REGION Network 6
   RUNG wire#powerrail
      Contact( #iStop )
      Contact( #iRun )
      wire#w1
      R_Coil( #oON )
   END_RUNG
   RUNG wire#powerrail
      Contact( #oBlocked )
   END_RUNG wire#w1
   RUNG wire#w1
      R_Coil( #oBrake )
   END_RUNG
   RUNG wire#w1
      R_Coil( #oContactor )
   END_RUNG
   // the same network as SCL:
   IF (#iStop AND #iRun) OR #oBlocked THEN
       #oON := FALSE;
       #oBrake := FALSE;
       #oContactor := FALSE;
   END_IF;
END_REGION

REGION Network 7
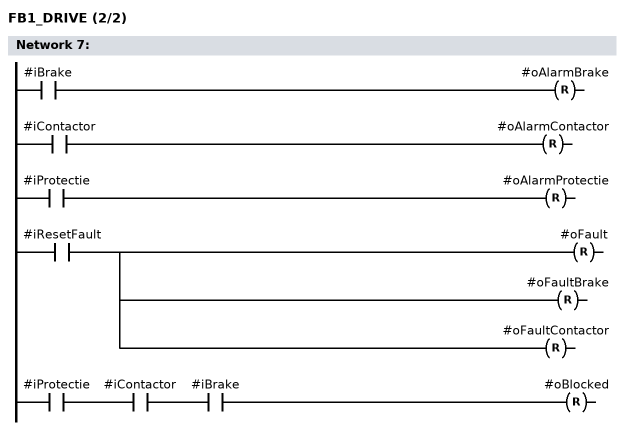
   RUNG wire#powerrail
      Contact( #iBrake )
      R_Coil( #oAlarmBrake )
   END_RUNG
   RUNG wire#powerrail
      Contact( #iContactor )
      R_Coil( #oAlarmContactor )
   END_RUNG
   RUNG wire#powerrail
      Contact( #iProtectie )
      R_Coil( #oAlarmProtectie )
   END_RUNG
   RUNG wire#powerrail
      Contact( #iResetFault )
      wire#w1
      R_Coil( #oFault )
   END_RUNG
   RUNG wire#w1
      R_Coil( #oFaultBrake )
   END_RUNG
   RUNG wire#w1
      R_Coil( #oFaultContactor )
   END_RUNG
   RUNG wire#powerrail
      Contact( #iProtectie )
      Contact( #iContactor )
      Contact( #iBrake )
      R_Coil( #oBlocked )
   END_RUNG
   // the same network as SCL:
   IF #iBrake THEN #oAlarmBrake := FALSE; END_IF;
   IF #iContactor THEN #oAlarmContactor := FALSE; END_IF;
   IF #iProtectie THEN #oAlarmProtectie := FALSE; END_IF;
   IF #iResetFault THEN
       #oFault := FALSE;
       #oFaultBrake := FALSE;
       #oFaultContactor := FALSE;
   END_IF;
   IF #iProtectie AND #iContactor AND #iBrake THEN #oBlocked := FALSE; END_IF;
END_REGION
END_FUNCTION_BLOCK

FUNCTION_BLOCK "FB_Pallet_Length"   // FB2, LAD
{ S7_Optimized_Access := 'TRUE' }
VERSION : 0.1
   VAR_INPUT
      iSQ_Pallet_Length : Bool;
      iConv_Speed : Int;
      Reset_Counter : Bool;
   END_VAR
   VAR_OUTPUT
      oPallet_Length : Int;
      oAlarm_Length : Bool;
   END_VAR
   VAR
      tSQ : Real;
      tMax : Time := T#20s;
      Pallet_count : Int;
      SQ_NOT : Bool;
      SQ_ON : Bool;
      Finished_counting : Bool;
   END_VAR
   VAR RETAIN
      Timer_ET : Time;
   END_VAR
   VAR
      Pallet_count_2 : Int;
      TON : TON_TIME;
   END_VAR
   VAR RETAIN
      CNT_PalletPass_2 : CTU_INT;
      CNT_PalletPass_1 : CTU_INT;
   END_VAR
   VAR_TEMP   // added for the SCL form of the ladder/FBD networks
      _w1 : Bool;
      _w2 : Bool;
   END_VAR
BEGIN

REGION Network 1
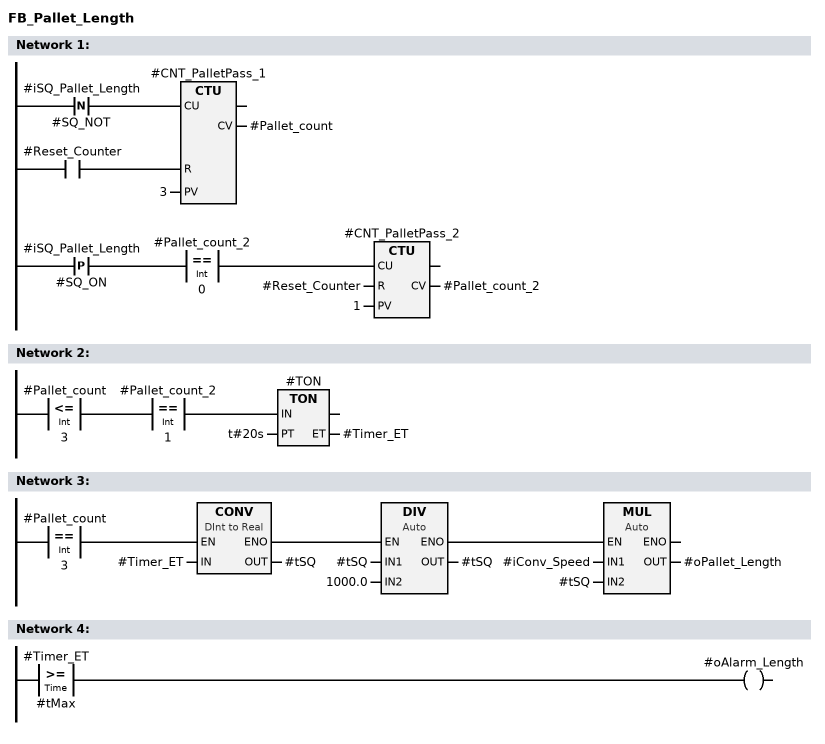
   #_w1 := NOT #iSQ_Pallet_Length AND #SQ_NOT;   // falling edge of #iSQ_Pallet_Length
   #SQ_NOT := #iSQ_Pallet_Length;
   #CNT_PalletPass_1(CU := #_w1, R := #Reset_Counter, PV := 3, CV => #Pallet_count);   // CTU
   #_w2 := #iSQ_Pallet_Length AND NOT #SQ_ON;   // rising edge of #iSQ_Pallet_Length
   #SQ_ON := #iSQ_Pallet_Length;
   #CNT_PalletPass_2(CU := #_w2 AND (#Pallet_count_2 = 0), R := #Reset_Counter, PV := 1, CV => #Pallet_count_2);   // CTU
END_REGION

REGION Network 2
   #TON(IN := (#Pallet_count <= 3) AND (#Pallet_count_2 = 1), PT := t#20s, ET => #Timer_ET);   // TON
END_REGION

REGION Network 3
   RUNG wire#powerrail
      { S7_Templates := "SrcType := Int" } EQ_Contact(in1 := #Pallet_count, in2 := 3)
      { S7_Templates := "[SrcType := DInt, DestType := Real]" } Convert(in := #Timer_ET, out => #tSQ)
      Div(in1 := #tSQ, in2 := 1000.0, out => #tSQ)
      Mul(in1 := #iConv_Speed, in2 := #tSQ, out => #oPallet_Length)
   END_RUNG
   // the same network as SCL:
   IF #Pallet_count = 3 THEN
       #tSQ := DINT_TO_REAL(#Timer_ET);
       #tSQ := #tSQ / 1000.0;
       #oPallet_Length := #iConv_Speed * #tSQ;
   END_IF;
END_REGION

REGION Network 4
   RUNG wire#powerrail
      { S7_Templates := "SrcType := Time" } GE_Contact(in1 := #Timer_ET, in2 := #tMax)
      Coil( #oAlarm_Length )
   END_RUNG
   // the same network as SCL:
   #oAlarm_Length := #Timer_ET >= #tMax;
END_REGION
END_FUNCTION_BLOCK

FUNCTION_BLOCK "FB_DS_Check_Machine"   // FB3, LAD
{ S7_Optimized_Access := 'TRUE' }
VERSION : 0.1
   VAR_INPUT
      iAir : Bool;
      iProtectie_CD_Drive : Bool;
      iProtectie_DS_Drive : Bool;
      iCD_Drive_Fault : Bool;
      iDS_Drive_Fault : Bool;
      iDestacker_Wait_Position : Bool;
      iSoftStarter_S1 : Bool;
      iSoftStarter_S2 : Bool;
   END_VAR
   VAR_OUTPUT
      oDS_Checked : Bool;
      oCD_Drive_NOK : Bool;
      oDS_Drive_NOK : Bool;
      oAir_NOK : Bool;
      oPower_NOK : Bool;
      oDestacker_NOK : Bool;
   END_VAR
   VAR
      AIR_OK : Bool;
      POWER_OK : Bool;
      Destacker_Wait_Position : Bool;
      CD_DRIVE_OK : Bool;
      DS_DRIVE_OK : Bool;
   END_VAR
BEGIN

REGION Network 1
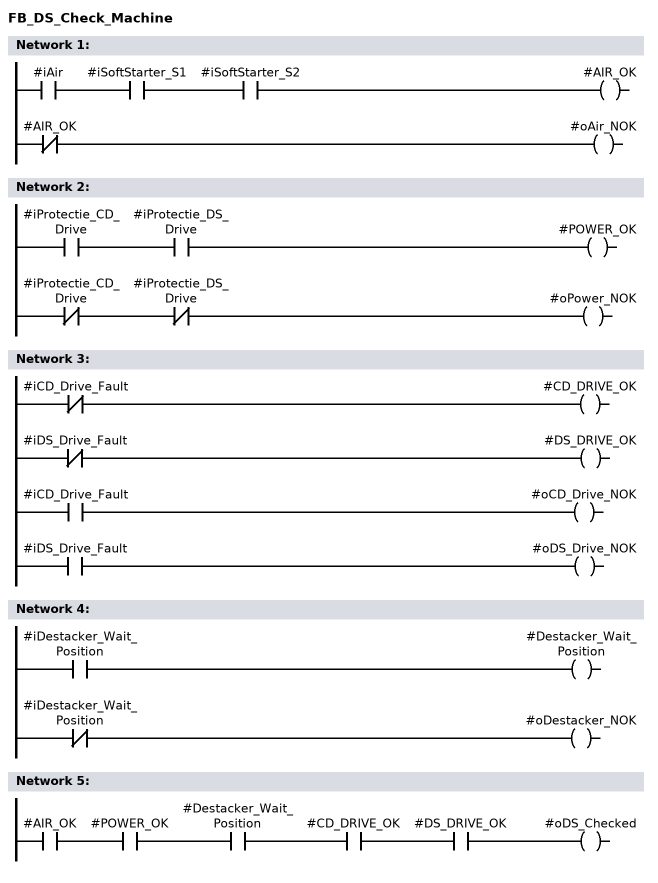
   RUNG wire#powerrail
      Contact( #iAir )
      Contact( #iSoftStarter_S1 )
      Contact( #iSoftStarter_S2 )
      Coil( #AIR_OK )
   END_RUNG
   RUNG wire#powerrail
      I_Contact( #AIR_OK )
      Coil( #oAir_NOK )
   END_RUNG
   // the same network as SCL:
   #AIR_OK := #iAir AND #iSoftStarter_S1 AND #iSoftStarter_S2;
   #oAir_NOK := NOT #AIR_OK;
END_REGION

REGION Network 2
   RUNG wire#powerrail
      Contact( #iProtectie_CD_Drive )
      Contact( #iProtectie_DS_Drive )
      Coil( #POWER_OK )
   END_RUNG
   RUNG wire#powerrail
      I_Contact( #iProtectie_CD_Drive )
      I_Contact( #iProtectie_DS_Drive )
      Coil( #oPower_NOK )
   END_RUNG
   // the same network as SCL:
   #POWER_OK := #iProtectie_CD_Drive AND #iProtectie_DS_Drive;
   #oPower_NOK := NOT #iProtectie_CD_Drive AND NOT #iProtectie_DS_Drive;
END_REGION

REGION Network 3
   RUNG wire#powerrail
      I_Contact( #iCD_Drive_Fault )
      Coil( #CD_DRIVE_OK )
   END_RUNG
   RUNG wire#powerrail
      I_Contact( #iDS_Drive_Fault )
      Coil( #DS_DRIVE_OK )
   END_RUNG
   RUNG wire#powerrail
      Contact( #iCD_Drive_Fault )
      Coil( #oCD_Drive_NOK )
   END_RUNG
   RUNG wire#powerrail
      Contact( #iDS_Drive_Fault )
      Coil( #oDS_Drive_NOK )
   END_RUNG
   // the same network as SCL:
   #CD_DRIVE_OK := NOT #iCD_Drive_Fault;
   #DS_DRIVE_OK := NOT #iDS_Drive_Fault;
   #oCD_Drive_NOK := #iCD_Drive_Fault;
   #oDS_Drive_NOK := #iDS_Drive_Fault;
END_REGION

REGION Network 4
   RUNG wire#powerrail
      Contact( #iDestacker_Wait_Position )
      Coil( #Destacker_Wait_Position )
   END_RUNG
   RUNG wire#powerrail
      I_Contact( #iDestacker_Wait_Position )
      Coil( #oDestacker_NOK )
   END_RUNG
   // the same network as SCL:
   #Destacker_Wait_Position := #iDestacker_Wait_Position;
   #oDestacker_NOK := NOT #iDestacker_Wait_Position;
END_REGION

REGION Network 5
   RUNG wire#powerrail
      Contact( #AIR_OK )
      Contact( #POWER_OK )
      Contact( #Destacker_Wait_Position )
      Contact( #CD_DRIVE_OK )
      Contact( #DS_DRIVE_OK )
      Coil( #oDS_Checked )
   END_RUNG
   // the same network as SCL:
   #oDS_Checked := #AIR_OK AND #POWER_OK AND #Destacker_Wait_Position AND #CD_DRIVE_OK AND #DS_DRIVE_OK;
END_REGION
END_FUNCTION_BLOCK

FUNCTION_BLOCK "FB_Init_S"   // FB4, LAD
TITLE = td -bitii de comenzi locali (ex: #Comanda_Furca) trebuie pusi in OUT
{ S7_Optimized_Access := 'TRUE' }
VERSION : 0.1
   VAR_INPUT
      DRV : "Bits_Stacker";
   END_VAR
   VAR
      Vertical : Bool;
      Furca : Bool;
      Comanda_Furca : Bool;
      Comanda_Vertical : Bool;
      InitReq : Bool;
      Init_OK : Bool;
      Alarm_Timeout_Vertical : Bool;
      Alarm_Timeout_Furca : Bool;
      "step" : USInt;
      Init_NotPossible : Bool;
      RstStack : Bool;
      Timer_Alarms : Array[0..1] of IEC_TIMER;
   END_VAR
   VAR_TEMP   // added for the SCL form of the ladder/FBD networks
      _w1 : Bool;
      _w2 : Bool;
   END_VAR
BEGIN

REGION Network 1: ini req
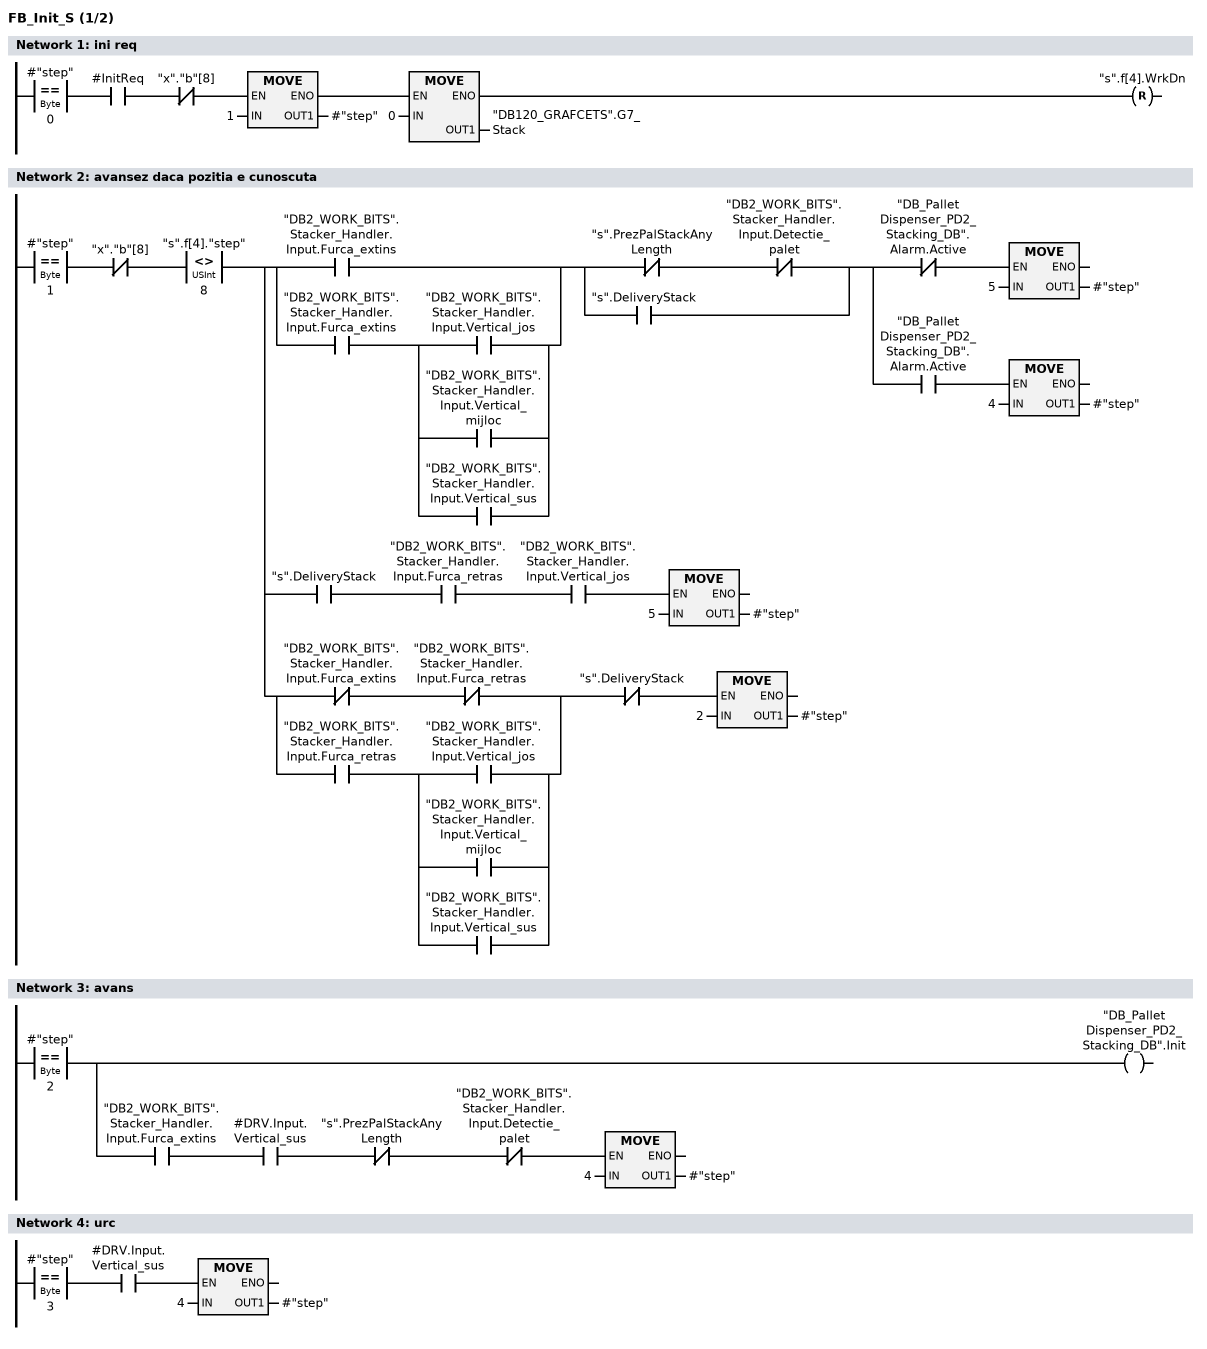
   RUNG wire#powerrail
      { S7_Templates := "SrcType := Byte" } EQ_Contact(in1 := #"step", in2 := 0)
      Contact( #InitReq )
      I_Contact( "x"."b"[8] )
      Move(in := 1, out1 => #"step")
      Move(in := 0, out1 => "DB120_GRAFCETS".G7_Stack)
      R_Coil( "s".f[4].WrkDn )
   END_RUNG
   // the same network as SCL:
   #_w1 := (#"step" = 0) AND #InitReq AND NOT "x"."b"[8];
   IF #_w1 THEN
       #"step" := 1;
       "DB120_GRAFCETS".G7_Stack := 0;
       "s".f[4].WrkDn := FALSE;
   END_IF;
END_REGION

REGION Network 2: avansez daca pozitia e cunoscuta
   RUNG wire#powerrail
      { S7_Templates := "SrcType := Byte" } EQ_Contact(in1 := #"step", in2 := 1)
      I_Contact( "x"."b"[8] )
      { S7_Templates := "SrcType := USInt" } NE_Contact(in1 := "s".f[4]."step", in2 := 8)
      wire#w1
      Contact( "DB2_WORK_BITS".Stacker_Handler.Input.Furca_extins )
      wire#w2
      I_Contact( "s".PrezPalStackAnyLength )
      I_Contact( "DB2_WORK_BITS".Stacker_Handler.Input.Detectie_palet )
      wire#w4
      I_Contact( "DB_PalletDispenser_PD2_Stacking_DB".Alarm.Active )
      Move(in := 5, out1 => #"step")
   END_RUNG
   RUNG wire#w1
      Contact( "DB2_WORK_BITS".Stacker_Handler.Input.Furca_extins )
      wire#w3
      Contact( "DB2_WORK_BITS".Stacker_Handler.Input.Vertical_jos )
   END_RUNG wire#w2
   RUNG wire#w3
      Contact( "DB2_WORK_BITS".Stacker_Handler.Input.Vertical_mijloc )
   END_RUNG wire#w2
   RUNG wire#w3
      Contact( "DB2_WORK_BITS".Stacker_Handler.Input.Vertical_sus )
   END_RUNG wire#w2
   RUNG wire#w2
      Contact( "s".DeliveryStack )
   END_RUNG wire#w4
   RUNG wire#w4
      Contact( "DB_PalletDispenser_PD2_Stacking_DB".Alarm.Active )
      Move(in := 4, out1 => #"step")
   END_RUNG
   RUNG wire#w1
      Contact( "s".DeliveryStack )
      Contact( "DB2_WORK_BITS".Stacker_Handler.Input.Furca_retras )
      Contact( "DB2_WORK_BITS".Stacker_Handler.Input.Vertical_jos )
      Move(in := 5, out1 => #"step")
   END_RUNG
   RUNG wire#w1
      I_Contact( "DB2_WORK_BITS".Stacker_Handler.Input.Furca_extins )
      I_Contact( "DB2_WORK_BITS".Stacker_Handler.Input.Furca_retras )
      wire#w5
      I_Contact( "s".DeliveryStack )
      Move(in := 2, out1 => #"step")
   END_RUNG
   RUNG wire#w1
      Contact( "DB2_WORK_BITS".Stacker_Handler.Input.Furca_retras )
      wire#w6
      Contact( "DB2_WORK_BITS".Stacker_Handler.Input.Vertical_jos )
   END_RUNG wire#w5
   RUNG wire#w6
      Contact( "DB2_WORK_BITS".Stacker_Handler.Input.Vertical_mijloc )
   END_RUNG wire#w5
   RUNG wire#w6
      Contact( "DB2_WORK_BITS".Stacker_Handler.Input.Vertical_sus )
   END_RUNG wire#w5
   // the same network as SCL:
   #_w1 := (#"step" = 1) AND NOT "x"."b"[8] AND ("s".f[4]."step" <> 8);
   #_w2 := #_w1 AND ("DB2_WORK_BITS".Stacker_Handler.Input.Furca_extins OR ("DB2_WORK_BITS".Stacker_Handler.Input.Furca_extins AND ("DB2_WORK_BITS".Stacker_Handler.Input.Vertical_jos OR "DB2_WORK_BITS".Stacker_Handler.Input.Vertical_mijloc OR "DB2_WORK_BITS".Stacker_Handler.Input.Vertical_sus))) AND ((NOT "s".PrezPalStackAnyLength AND NOT "DB2_WORK_BITS".Stacker_Handler.Input.Detectie_palet) OR "s".DeliveryStack);
   IF #_w2 AND NOT "DB_PalletDispenser_PD2_Stacking_DB".Alarm.Active THEN #"step" := 5; END_IF;
   IF #_w2 AND "DB_PalletDispenser_PD2_Stacking_DB".Alarm.Active THEN #"step" := 4; END_IF;
   IF #_w1 AND "s".DeliveryStack AND "DB2_WORK_BITS".Stacker_Handler.Input.Furca_retras AND "DB2_WORK_BITS".Stacker_Handler.Input.Vertical_jos THEN
       #"step" := 5;
   END_IF;
   IF #_w1 AND ((NOT "DB2_WORK_BITS".Stacker_Handler.Input.Furca_extins AND NOT "DB2_WORK_BITS".Stacker_Handler.Input.Furca_retras) OR ("DB2_WORK_BITS".Stacker_Handler.Input.Furca_retras AND ("DB2_WORK_BITS".Stacker_Handler.Input.Vertical_jos OR "DB2_WORK_BITS".Stacker_Handler.Input.Vertical_mijloc OR "DB2_WORK_BITS".Stacker_Handler.Input.Vertical_sus))) AND NOT "s".DeliveryStack THEN
       #"step" := 2;
   END_IF;
END_REGION

REGION Network 3: avans
   RUNG wire#powerrail
      { S7_Templates := "SrcType := Byte" } EQ_Contact(in1 := #"step", in2 := 2)
      wire#w1
      Coil( "DB_PalletDispenser_PD2_Stacking_DB".Init )
   END_RUNG
   RUNG wire#w1
      Contact( "DB2_WORK_BITS".Stacker_Handler.Input.Furca_extins )
      Contact( #DRV.Input.Vertical_sus )
      I_Contact( "s".PrezPalStackAnyLength )
      I_Contact( "DB2_WORK_BITS".Stacker_Handler.Input.Detectie_palet )
      Move(in := 4, out1 => #"step")
   END_RUNG
   // the same network as SCL:
   "DB_PalletDispenser_PD2_Stacking_DB".Init := #"step" = 2;
   IF "DB_PalletDispenser_PD2_Stacking_DB".Init AND "DB2_WORK_BITS".Stacker_Handler.Input.Furca_extins AND #DRV.Input.Vertical_sus AND NOT "s".PrezPalStackAnyLength AND NOT "DB2_WORK_BITS".Stacker_Handler.Input.Detectie_palet THEN
       #"step" := 4;
   END_IF;
END_REGION

REGION Network 4: urc
   RUNG wire#powerrail
      { S7_Templates := "SrcType := Byte" } EQ_Contact(in1 := #"step", in2 := 3)
      Contact( #DRV.Input.Vertical_sus )
      Move(in := 4, out1 => #"step")
   END_RUNG
   // the same network as SCL:
   IF (#"step" = 3) AND #DRV.Input.Vertical_sus THEN #"step" := 4; END_IF;
END_REGION

REGION Network 5: Reset FB stacker errors
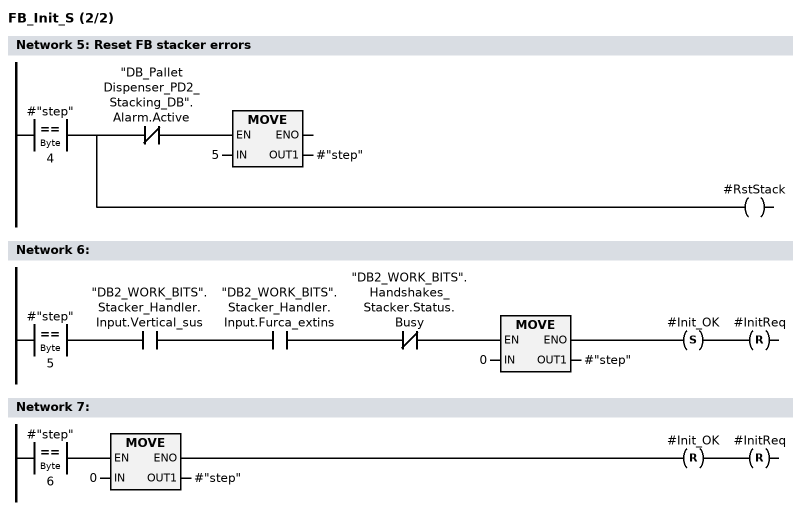
   RUNG wire#powerrail
      { S7_Templates := "SrcType := Byte" } EQ_Contact(in1 := #"step", in2 := 4)
      wire#w1
      I_Contact( "DB_PalletDispenser_PD2_Stacking_DB".Alarm.Active )
      Move(in := 5, out1 => #"step")
   END_RUNG
   RUNG wire#w1
      Coil( #RstStack )
   END_RUNG
   // the same network as SCL:
   #_w1 := #"step" = 4;
   IF #_w1 AND NOT "DB_PalletDispenser_PD2_Stacking_DB".Alarm.Active THEN #"step" := 5; END_IF;
   #RstStack := #_w1;
END_REGION

REGION Network 6
   RUNG wire#powerrail
      { S7_Templates := "SrcType := Byte" } EQ_Contact(in1 := #"step", in2 := 5)
      Contact( "DB2_WORK_BITS".Stacker_Handler.Input.Vertical_sus )
      Contact( "DB2_WORK_BITS".Stacker_Handler.Input.Furca_extins )
      I_Contact( "DB2_WORK_BITS".Handshakes_Stacker.Status.Busy )
      Move(in := 0, out1 => #"step")
      S_Coil( #Init_OK )
      R_Coil( #InitReq )
   END_RUNG
   // the same network as SCL:
   #_w1 := (#"step" = 5) AND "DB2_WORK_BITS".Stacker_Handler.Input.Vertical_sus AND "DB2_WORK_BITS".Stacker_Handler.Input.Furca_extins AND NOT "DB2_WORK_BITS".Handshakes_Stacker.Status.Busy;
   IF #_w1 THEN
       #"step" := 0;
       #Init_OK := TRUE;
       #InitReq := FALSE;
   END_IF;
END_REGION

REGION Network 7
   RUNG wire#powerrail
      { S7_Templates := "SrcType := Byte" } EQ_Contact(in1 := #"step", in2 := 6)
      Move(in := 0, out1 => #"step")
      R_Coil( #Init_OK )
      R_Coil( #InitReq )
   END_RUNG
   // the same network as SCL:
   #_w1 := #"step" = 6;
   IF #_w1 THEN
       #"step" := 0;
       #Init_OK := FALSE;
       #InitReq := FALSE;
   END_IF;
END_REGION
END_FUNCTION_BLOCK

FUNCTION_BLOCK "FB_Centrare"   // FB5, LAD
{ S7_Optimized_Access := 'TRUE' }
VERSION : 0.1
   VAR_INPUT
      Senzor_eliber : Bool;
      senzor_centr : Bool;
      step_st : USInt;
   END_VAR
   VAR_OUTPUT
      Comanda_centr : Bool;
      Comanda_eliber : Bool;
      stpo : USInt;
   END_VAR
   VAR_IN_OUT
      work : Bool;
   END_VAR
   VAR
      "step" : USInt;
      cmdav : Bool;
      cmdret : Bool;
      tmr : Array[1..3] of IEC_TIMER;
   END_VAR
   VAR_TEMP   // added for the SCL form of the ladder/FBD networks
      _w1 : Bool;
      _w2 : Bool;
   END_VAR
BEGIN

REGION Network 1
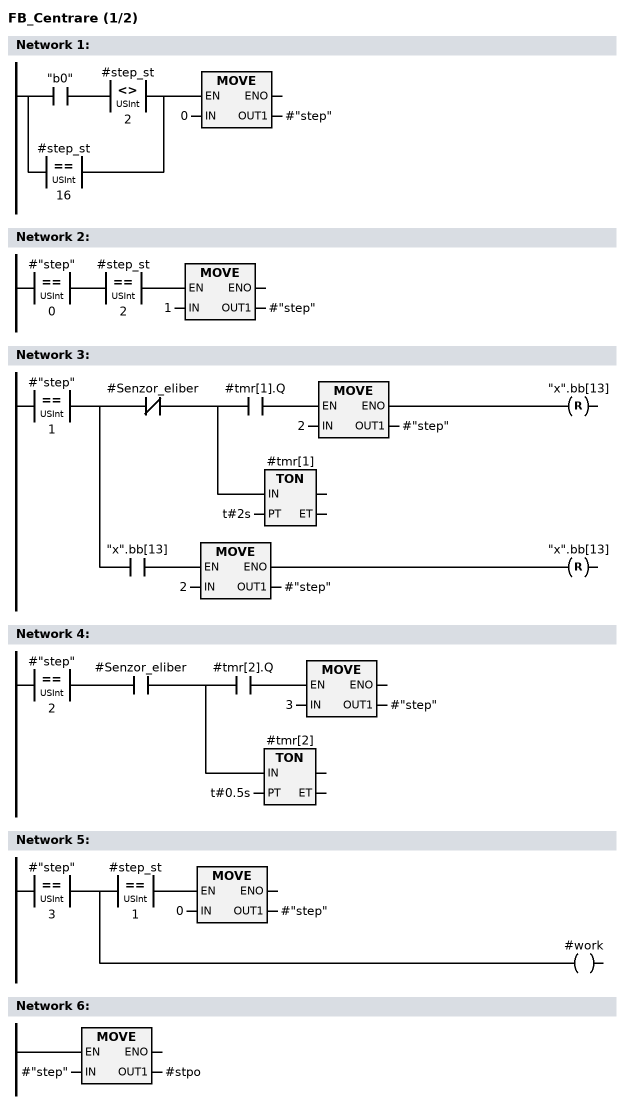
   RUNG wire#powerrail
      Contact( "b0" )
      { S7_Templates := "SrcType := USInt" } NE_Contact(in1 := #step_st, in2 := 2)
      wire#w1
      Move(in := 0, out1 => #"step")
   END_RUNG
   RUNG wire#powerrail
      { S7_Templates := "SrcType := USInt" } EQ_Contact(in1 := #step_st, in2 := 16)
   END_RUNG wire#w1
   // the same network as SCL:
   IF ("b0" AND (#step_st <> 2)) OR (#step_st = 16) THEN #"step" := 0; END_IF;
END_REGION

REGION Network 2
   RUNG wire#powerrail
      { S7_Templates := "SrcType := USInt" } EQ_Contact(in1 := #"step", in2 := 0)
      { S7_Templates := "SrcType := USInt" } EQ_Contact(in1 := #step_st, in2 := 2)
      Move(in := 1, out1 => #"step")
   END_RUNG
   // the same network as SCL:
   IF (#"step" = 0) AND (#step_st = 2) THEN #"step" := 1; END_IF;
END_REGION

REGION Network 3
   #_w1 := #"step" = 1;
   #_w2 := #_w1 AND NOT #Senzor_eliber;
   IF #_w2 AND #tmr[1].Q THEN
       #"step" := 2;
       "x".bb[13] := FALSE;
   END_IF;
   #tmr[1].TON(IN := #_w2, PT := t#2s);
   IF #_w1 AND "x".bb[13] THEN
       #"step" := 2;
       "x".bb[13] := FALSE;
   END_IF;
END_REGION

REGION Network 4
   #_w1 := (#"step" = 2) AND #Senzor_eliber;
   IF #_w1 AND #tmr[2].Q THEN #"step" := 3; END_IF;
   #tmr[2].TON(IN := #_w1, PT := t#0.5s);
END_REGION

REGION Network 5
   RUNG wire#powerrail
      { S7_Templates := "SrcType := USInt" } EQ_Contact(in1 := #"step", in2 := 3)
      wire#w1
      { S7_Templates := "SrcType := USInt" } EQ_Contact(in1 := #step_st, in2 := 1)
      Move(in := 0, out1 => #"step")
   END_RUNG
   RUNG wire#w1
      Coil( #work )
   END_RUNG
   // the same network as SCL:
   #_w1 := #"step" = 3;
   IF #_w1 AND (#step_st = 1) THEN #"step" := 0; END_IF;
   #work := #_w1;
END_REGION

REGION Network 6
   RUNG wire#powerrail
      Move(in := #"step", out1 => #stpo)
   END_RUNG
   // the same network as SCL:
   #stpo := #"step";
END_REGION

REGION Network 7: Apelare centror
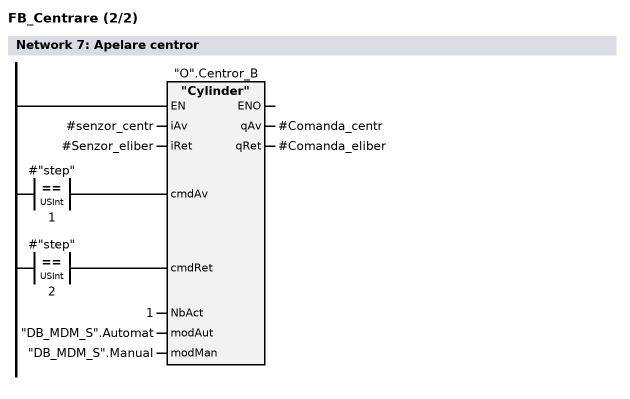
   RUNG wire#powerrail
      "O".Centror_B(cmdAv := wire#w1, cmdRet := wire#w2, iAv := #senzor_centr, iRet := #Senzor_eliber, NbAct := 1, modAut := "DB_MDM_S".Automat, modMan := "DB_MDM_S".Manual, qAv => #Comanda_centr, qRet => #Comanda_eliber)
   END_RUNG
   RUNG wire#powerrail
      { S7_Templates := "SrcType := USInt" } EQ_Contact(in1 := #"step", in2 := 1)
   END_RUNG wire#w1
   RUNG wire#powerrail
      { S7_Templates := "SrcType := USInt" } EQ_Contact(in1 := #"step", in2 := 2)
   END_RUNG wire#w2
   // the same network as SCL:
   "O".Centror_B(iAv := #senzor_centr,   // "Cylinder"
                 iRet := #Senzor_eliber,
                 cmdAv := #"step" = 1,
                 cmdRet := #"step" = 2,
                 NbAct := 1,
                 modAut := "DB_MDM_S".Automat,
                 modMan := "DB_MDM_S".Manual,
                 qAv => #Comanda_centr,
                 qRet => #Comanda_eliber);
END_REGION
END_FUNCTION_BLOCK

FUNCTION_BLOCK "sim"   // FB6, LAD
{ S7_Optimized_Access := 'TRUE' }
VERSION : 0.1
   VAR
      cen : "simCylinder";
      stH : "simCylinder";
      tct : IEC_TIMER;
      tct2 : Bool;
      tct1 : Bool;
      tm : Array[0..10] of IEC_TIMER;
      "Prezenta palet_dreapta" : Bool;
   END_VAR
   VAR_TEMP   // added for the SCL form of the ladder/FBD networks
      _w1 : Bool;
      _w2 : Bool;
   END_VAR
BEGIN

REGION Network 1
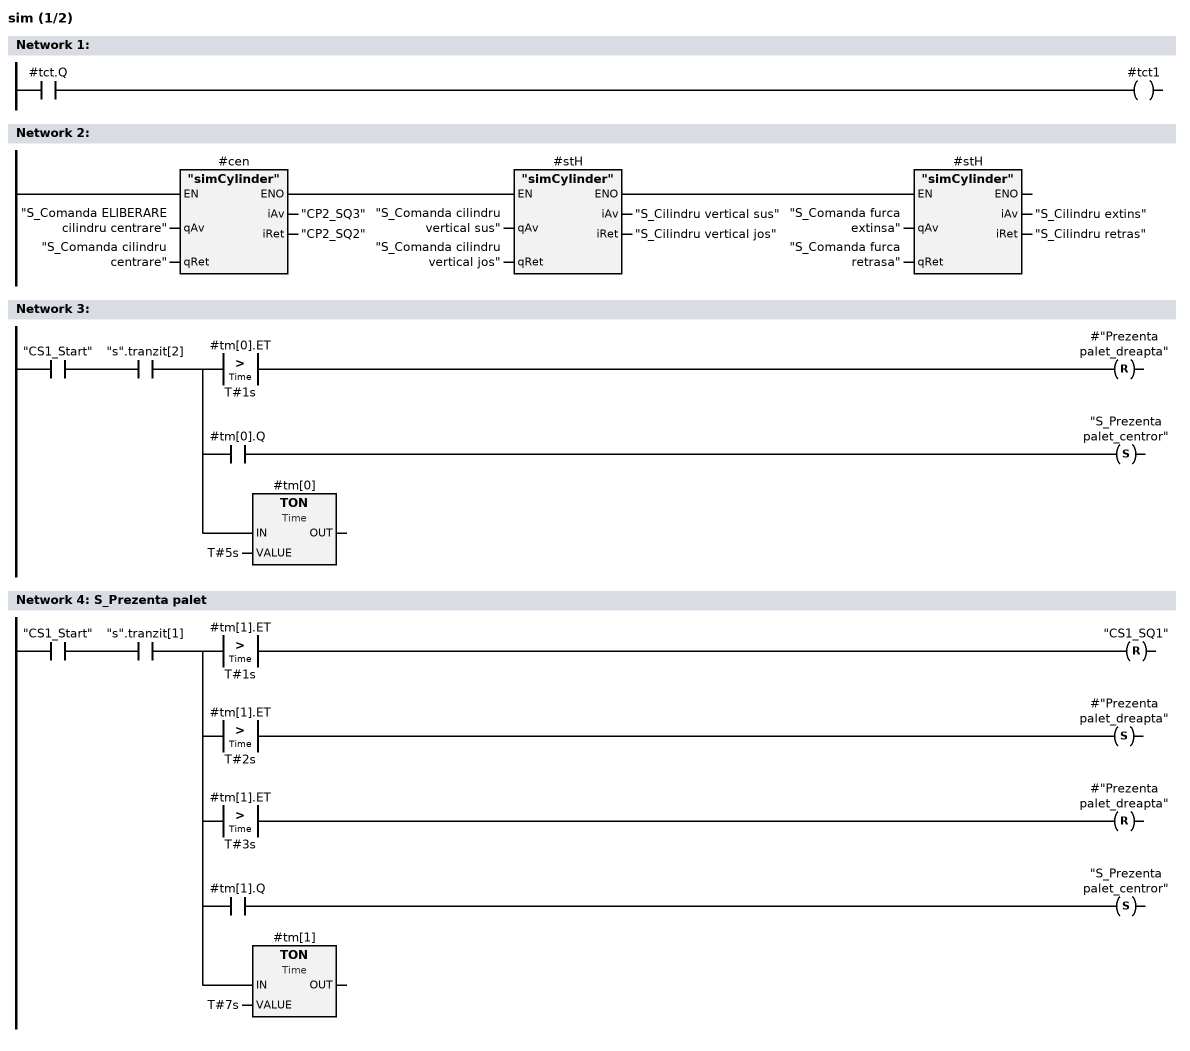
   RUNG wire#powerrail
      Contact( #tct.Q )
      Coil( #tct1 )
   END_RUNG
   // the same network as SCL:
   #tct1 := #tct.Q;
END_REGION

REGION Network 2
   RUNG wire#powerrail
      #cen(qAv := "S_Comanda ELIBERARE cilindru centrare", qRet := "S_Comanda cilindru centrare", iAv => "CP2_SQ3", iRet => "CP2_SQ2")
      #stH(qAv := "S_Comanda cilindru vertical sus", qRet := "S_Comanda cilindru vertical jos", iAv => "S_Cilindru vertical sus", iRet => "S_Cilindru vertical jos")
      #stH(qAv := "S_Comanda furca extinsa", qRet := "S_Comanda furca retrasa", iAv => "S_Cilindru extins", iRet => "S_Cilindru retras")
   END_RUNG
   // the same network as SCL:
   #cen(qAv := "S_Comanda ELIBERARE cilindru centrare",   // "simCylinder"
        qRet := "S_Comanda cilindru centrare",
        iAv => "CP2_SQ3",
        iRet => "CP2_SQ2",
        ENO => #_w1);
   #stH(EN := #_w1,   // "simCylinder"
        qAv := "S_Comanda cilindru vertical sus",
        qRet := "S_Comanda cilindru vertical jos",
        iAv => "S_Cilindru vertical sus",
        iRet => "S_Cilindru vertical jos",
        ENO => #_w2);
   IF #_w2 THEN
       #stH(qAv := "S_Comanda furca extinsa",   // "simCylinder"
            qRet := "S_Comanda furca retrasa",
            iAv => "S_Cilindru extins",
            iRet => "S_Cilindru retras");
   END_IF;
END_REGION

REGION Network 3
   #_w1 := "CS1_Start" AND "s".tranzit[2];
   IF #_w1 AND (#tm[0].ET > T#1s) THEN #"Prezenta palet_dreapta" := FALSE; END_IF;
   IF #_w1 AND #tm[0].Q THEN "S_Prezenta palet_centror" := TRUE; END_IF;
   #tm[0].TON(IN := #_w1, PT := T#5s);   // TON coil
END_REGION

REGION Network 4: S_Prezenta palet
   #_w1 := "CS1_Start" AND "s".tranzit[1];
   IF #_w1 AND (#tm[1].ET > T#1s) THEN "CS1_SQ1" := FALSE; END_IF;
   IF #_w1 AND (#tm[1].ET > T#2s) THEN #"Prezenta palet_dreapta" := TRUE; END_IF;
   IF #_w1 AND (#tm[1].ET > T#3s) THEN #"Prezenta palet_dreapta" := FALSE; END_IF;
   IF #_w1 AND #tm[1].Q THEN "S_Prezenta palet_centror" := TRUE; END_IF;
   #tm[1].TON(IN := #_w1, PT := T#7s);   // TON coil
END_REGION

REGION Network 5
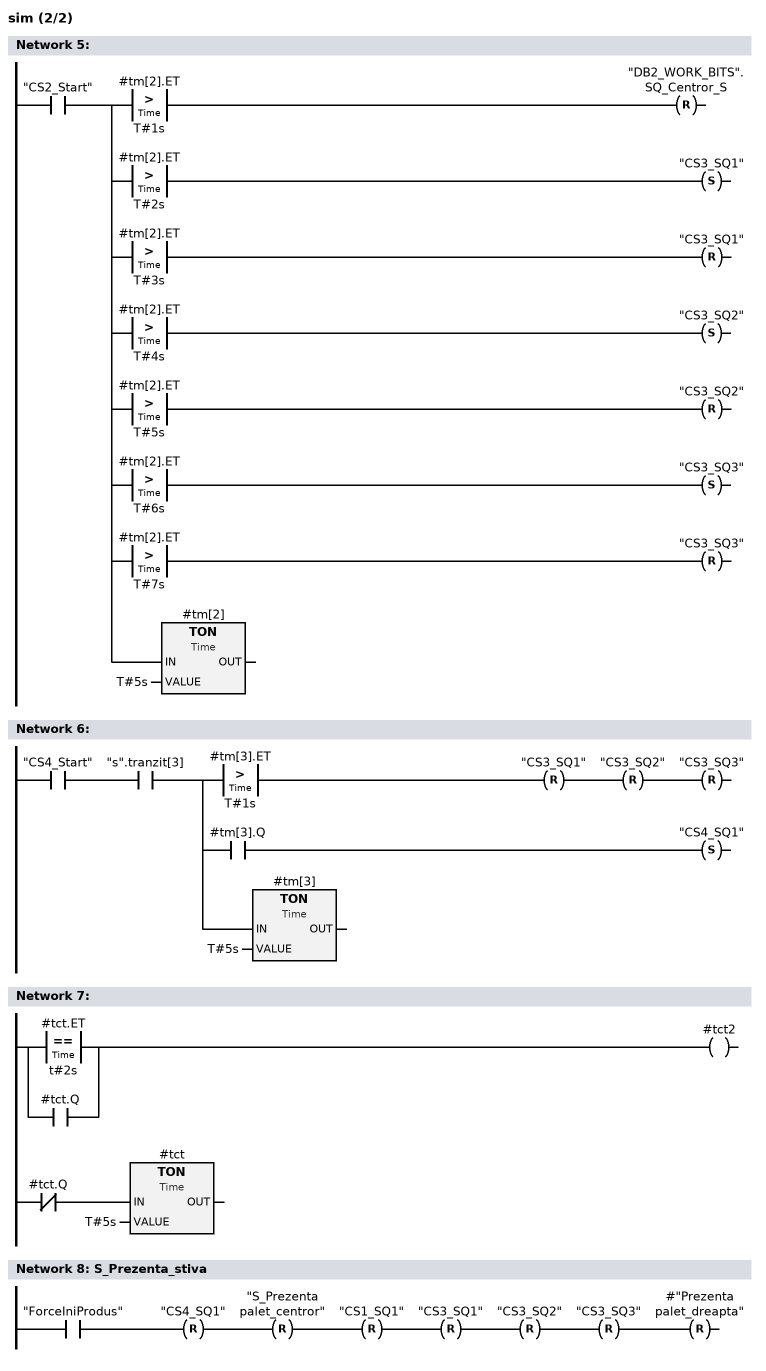
   IF "CS2_Start" AND (#tm[2].ET > T#1s) THEN "DB2_WORK_BITS".SQ_Centror_S := FALSE; END_IF;
   IF "CS2_Start" AND (#tm[2].ET > T#2s) THEN "CS3_SQ1" := TRUE; END_IF;
   IF "CS2_Start" AND (#tm[2].ET > T#3s) THEN "CS3_SQ1" := FALSE; END_IF;
   IF "CS2_Start" AND (#tm[2].ET > T#4s) THEN "CS3_SQ2" := TRUE; END_IF;
   IF "CS2_Start" AND (#tm[2].ET > T#5s) THEN "CS3_SQ2" := FALSE; END_IF;
   IF "CS2_Start" AND (#tm[2].ET > T#6s) THEN "CS3_SQ3" := TRUE; END_IF;
   IF "CS2_Start" AND (#tm[2].ET > T#7s) THEN "CS3_SQ3" := FALSE; END_IF;
   #tm[2].TON(IN := "CS2_Start", PT := T#5s);   // TON coil
END_REGION

REGION Network 6
   #_w1 := "CS4_Start" AND "s".tranzit[3];
   IF #_w1 AND (#tm[3].ET > T#1s) THEN
       "CS3_SQ1" := FALSE;
       "CS3_SQ2" := FALSE;
       "CS3_SQ3" := FALSE;
   END_IF;
   IF #_w1 AND #tm[3].Q THEN "CS4_SQ1" := TRUE; END_IF;
   #tm[3].TON(IN := #_w1, PT := T#5s);   // TON coil
END_REGION

REGION Network 7
   #tct2 := (#tct.ET = t#2s) OR #tct.Q;
   #tct.TON(IN := NOT #tct.Q, PT := T#5s);   // TON coil
END_REGION

REGION Network 8: S_Prezenta_stiva
   RUNG wire#powerrail
      Contact( "ForceIniProdus" )
      R_Coil( "CS4_SQ1" )
      R_Coil( "S_Prezenta palet_centror" )
      R_Coil( "CS1_SQ1" )
      R_Coil( "CS3_SQ1" )
      R_Coil( "CS3_SQ2" )
      R_Coil( "CS3_SQ3" )
      R_Coil( #"Prezenta palet_dreapta" )
   END_RUNG
   // the same network as SCL:
   IF "ForceIniProdus" THEN
       "CS4_SQ1" := FALSE;
       "S_Prezenta palet_centror" := FALSE;
       "CS1_SQ1" := FALSE;
       "CS3_SQ1" := FALSE;
       "CS3_SQ2" := FALSE;
       "CS3_SQ3" := FALSE;
       #"Prezenta palet_dreapta" := FALSE;
   END_IF;
END_REGION
END_FUNCTION_BLOCK

FUNCTION_BLOCK "Cylinder"   // FB7, LAD
{ S7_Optimized_Access := 'TRUE' }
VERSION : 0.1
   VAR_INPUT
      iAv : Bool;
      iRet : Bool;
      cmdAv : Bool;
      cmdRet : Bool;
      NbAct : SInt;
      modAut : Bool;
      modMan : Bool;
   END_VAR
   VAR_OUTPUT
      qAv : Bool;
      qRet : Bool;
   END_VAR
   VAR
      tmrAv : IEC_TIMER;
      tmrRet : IEC_TIMER;
      tmrLoseAv : IEC_TIMER;
      tmrLoseRet : IEC_TIMER;
      tmrNoReleaseAv : IEC_TIMER;
      tmrNoReleaseRet : IEC_TIMER;
      tmrDelayAv : IEC_TIMER;
      tmrDelayRet : IEC_TIMER;
      memAv : Bool;
      memRet : Bool;
      almTmtAv : Bool;
      almTmtRet : Bool;
      almLoseAv : Bool;
      almLoseRet : Bool;
      almNoReleaseAv : Bool;
      almNoReleaseRet : Bool;
      almDiscordance : Bool;
      alm : Bool;
      HMI_stat : SInt;
      EnAv : Bool;
      EnRet : Bool;
      ButAv : Bool;
      ButRet : Bool;
      StatAv : USInt;
      StatRet : USInt;
      AlarmW : Word;
      tr : USInt;
   END_VAR
   VAR CONSTANT
      b0 : Bool;
   END_VAR
   VAR_TEMP   // added for the SCL form of the ladder/FBD networks
      _w1 : Bool;
   END_VAR
BEGIN

REGION Network 1: memorii stare pt alarma de disparitie
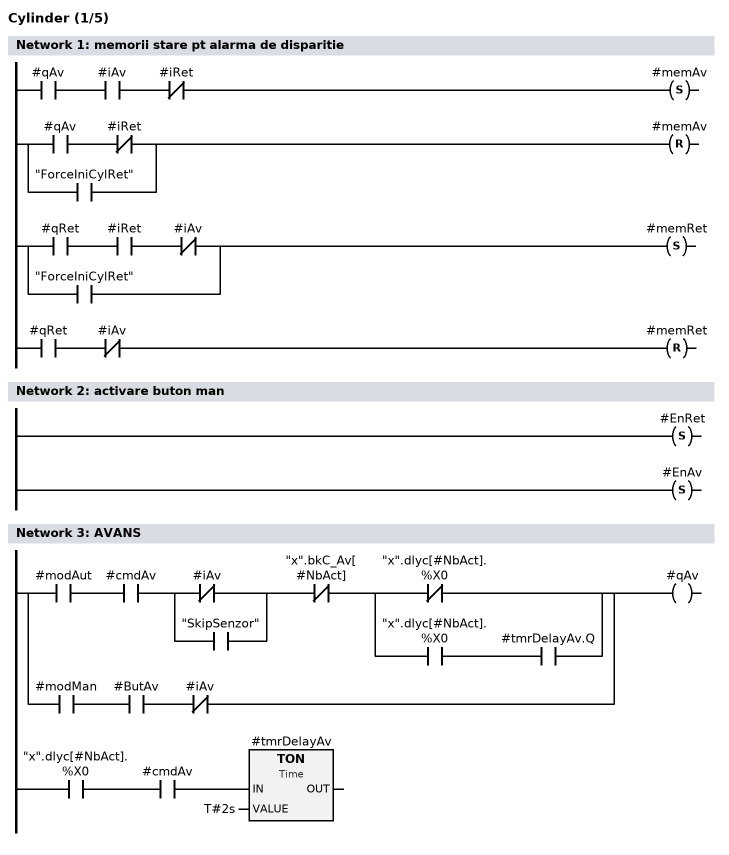
   RUNG wire#powerrail
      Contact( #qAv )
      Contact( #iAv )
      I_Contact( #iRet )
      S_Coil( #memAv )
   END_RUNG
   RUNG wire#powerrail
      Contact( #qAv )
      I_Contact( #iRet )
      wire#w1
      R_Coil( #memAv )
   END_RUNG
   RUNG wire#powerrail
      Contact( "ForceIniCylRet" )
   END_RUNG wire#w1
   RUNG wire#powerrail
      Contact( #qRet )
      Contact( #iRet )
      I_Contact( #iAv )
      wire#w2
      S_Coil( #memRet )
   END_RUNG
   RUNG wire#powerrail
      Contact( "ForceIniCylRet" )
   END_RUNG wire#w2
   RUNG wire#powerrail
      Contact( #qRet )
      I_Contact( #iAv )
      R_Coil( #memRet )
   END_RUNG
   // the same network as SCL:
   IF #qAv AND #iAv AND NOT #iRet THEN #memAv := TRUE; END_IF;
   IF (#qAv AND NOT #iRet) OR "ForceIniCylRet" THEN #memAv := FALSE; END_IF;
   IF (#qRet AND #iRet AND NOT #iAv) OR "ForceIniCylRet" THEN #memRet := TRUE; END_IF;
   IF #qRet AND NOT #iAv THEN #memRet := FALSE; END_IF;
END_REGION

REGION Network 2: activare buton man
   RUNG wire#powerrail
      S_Coil( #EnRet )
   END_RUNG
   RUNG wire#powerrail
      S_Coil( #EnAv )
   END_RUNG
   // the same network as SCL:
   #EnRet := TRUE;
   #EnAv := TRUE;
END_REGION

REGION Network 3: AVANS
   #qAv := (#modAut AND #cmdAv AND (NOT #iAv OR "SkipSenzor") AND NOT "x".bkC_Av[#NbAct] AND (NOT "x".dlyc[#NbAct].%X0 OR ("x".dlyc[#NbAct].%X0 AND #tmrDelayAv.Q))) OR (#modMan AND #ButAv AND NOT #iAv);
   #tmrDelayAv.TON(IN := "x".dlyc[#NbAct].%X0 AND #cmdAv, PT := T#2s);   // TON coil
END_REGION

REGION Network 4: trace
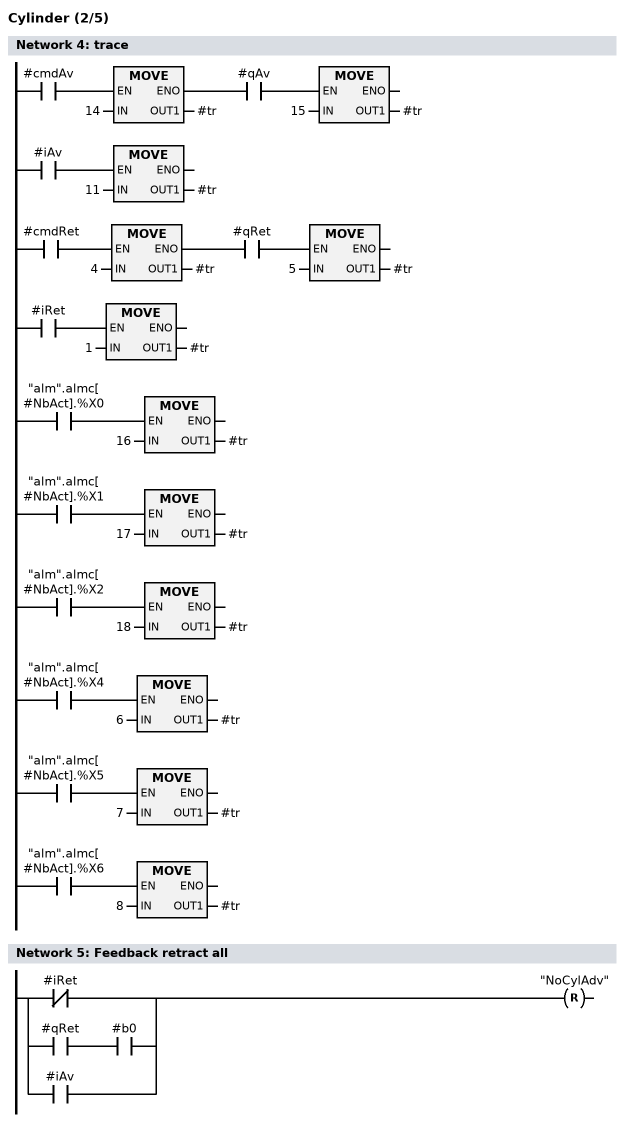
   RUNG wire#powerrail
      Contact( #cmdAv )
      Move(in := 14, out1 => #tr)
      Contact( #qAv )
      Move(in := 15, out1 => #tr)
   END_RUNG
   RUNG wire#powerrail
      Contact( #iAv )
      Move(in := 11, out1 => #tr)
   END_RUNG
   RUNG wire#powerrail
      Contact( #cmdRet )
      Move(in := 4, out1 => #tr)
      Contact( #qRet )
      Move(in := 5, out1 => #tr)
   END_RUNG
   RUNG wire#powerrail
      Contact( #iRet )
      Move(in := 1, out1 => #tr)
   END_RUNG
   RUNG wire#powerrail
      Contact( "alm".almc[#NbAct].%X0 )
      Move(in := 16, out1 => #tr)
   END_RUNG
   RUNG wire#powerrail
      Contact( "alm".almc[#NbAct].%X1 )
      Move(in := 17, out1 => #tr)
   END_RUNG
   RUNG wire#powerrail
      Contact( "alm".almc[#NbAct].%X2 )
      Move(in := 18, out1 => #tr)
   END_RUNG
   RUNG wire#powerrail
      Contact( "alm".almc[#NbAct].%X4 )
      Move(in := 6, out1 => #tr)
   END_RUNG
   RUNG wire#powerrail
      Contact( "alm".almc[#NbAct].%X5 )
      Move(in := 7, out1 => #tr)
   END_RUNG
   RUNG wire#powerrail
      Contact( "alm".almc[#NbAct].%X6 )
      Move(in := 8, out1 => #tr)
   END_RUNG
   // the same network as SCL:
   IF #cmdAv THEN #tr := 14; END_IF;
   IF #cmdAv AND #qAv THEN #tr := 15; END_IF;
   IF #iAv THEN #tr := 11; END_IF;
   IF #cmdRet THEN #tr := 4; END_IF;
   IF #cmdRet AND #qRet THEN #tr := 5; END_IF;
   IF #iRet THEN #tr := 1; END_IF;
   IF "alm".almc[#NbAct].%X0 THEN #tr := 16; END_IF;
   IF "alm".almc[#NbAct].%X1 THEN #tr := 17; END_IF;
   IF "alm".almc[#NbAct].%X2 THEN #tr := 18; END_IF;
   IF "alm".almc[#NbAct].%X4 THEN #tr := 6; END_IF;
   IF "alm".almc[#NbAct].%X5 THEN #tr := 7; END_IF;
   IF "alm".almc[#NbAct].%X6 THEN #tr := 8; END_IF;
END_REGION

REGION Network 5: Feedback retract all
   RUNG wire#powerrail
      I_Contact( #iRet )
      wire#w1
      R_Coil( "NoCylAdv" )
   END_RUNG
   RUNG wire#powerrail
      Contact( #qRet )
      Contact( #b0 )
   END_RUNG wire#w1
   RUNG wire#powerrail
      Contact( #iAv )
   END_RUNG wire#w1
   // the same network as SCL:
   IF NOT #iRet OR (#qRet AND #b0) OR #iAv THEN "NoCylAdv" := FALSE; END_IF;
END_REGION

REGION Network 6: RETRAG